        [6].Andco_Values.Pounds_Per_Inch := 65.0, [6].Andco_Values.New_Rate := 4000.0, [6].Andco_Values.Analog := 1, [6].Andco_Values.Min_Position := 625, [6].Andco_Values.Length := 12.0, [6].Andco_Values.InchesOpen := 7.1282053, [6].Andco_Values.AnalogValue := 9660, [6].Clean_Load_Delay_Stop := 36000, [6].Treat_Load_Delay_Stop := 34000, [6].tmrStopDelay.EN := 1, [6].tmrStopDelay.TT := 1, [6].Available_For_Clean_Load := 1, [6].Available_For_Treat_Load := 1, [7].Bin_Description := '10', [7].Bin_Variety.Item_Number := '823001', [7].Bin_Variety.Name := 'ARTDECO CERTIFIED FALL SWH', [7].Bin_Variety.Class := 'Certified', [7].Bin_Variety.Color[0].Color := 1, [7].Rate_Cal_Points[1].Andco_Position := 3007, [7].Rate_Cal_Points[1].Rate := 1000, [7].Rate_Cal_Points[2].Andco_Position := 5443, [7].Rate_Cal_Points[2].Rate := 2000, [7].Rate_Cal_Points[3].Andco_Position := 7342, [7].Rate_Cal_Points[3].Rate := 3000, [7].Rate_Cal_Points[4].Andco_Position := 9304, [7].Rate_Cal_Points[4].Rate := 4000, [7].Clean_Load_Delay_Start := 36500, [7].Treat_Load_Delay_Start := 30000, [7].Andco_Values.Cal_Status := 4, [7].Andco_Values.Raw_Position := 9878, [7].Andco_Values.Max_Position := 10246, [7].Andco_Values.Preact := 20, [7].Andco_Values.Percent_Open := 0.9646484, [7].Andco_Values.New_Pos := 68, [7].Andco_Values.Width := 6.0, [7].Andco_Values.Rate := 4292.5586, [7].Andco_Values.Pounds_Per_Inch := 65.0, [7].Andco_Values.New_Rate := 3700.0, [7].Andco_Values.Analog := 1, [7].Andco_Values.Min_Position := 6, [7].Andco_Values.Length := 12.0, [7].Andco_Values.InchesOpen := 11.575781, [7].Andco_Values.AnalogValue := 9884, [7].Clean_Load_Delay_Stop := 36500, [7].Treat_Load_Delay_Stop := 33000, [7].tmrStopDelay.EN := 1, [7].tmrStopDelay.TT := 1, [7].Available_For_Clean_Load := 1, [7].Available_For_Treat_Load := 1, [8].Bin_Description := '12', [8].Bin_Variety.Name := 'Empty', [8].Bin_Variety.Color[0].Color := 1, [8].Rate_Cal_Points[1].Andco_Position := 3358, [8].Rate_Cal_Points[1].Rate := 1000, [8].Rate_Cal_Points[2].Andco_Position := 5110, [8].Rate_Cal_Points[2].Rate := 2000, [8].Rate_Cal_Points[3].Andco_Position := 6534, [8].Rate_Cal_Points[3].Rate := 3000, [8].Rate_Cal_Points[4].Andco_Position := 8210, [8].Rate_Cal_Points[4].Rate := 4000,
        [8].Clean_Load_Delay_Start := 37000, [8].Treat_Load_Delay_Start := 31000, [8].Andco_Values.Cal_Status := 4, [8].Andco_Values.Raw_Position := 8474, [8].Andco_Values.Max_Position := 15055, [8].Andco_Values.Preact := 20, [8].Andco_Values.Percent_Open := 0.66141117, [8].Andco_Values.New_Pos := 61, [8].Andco_Values.Width := 6.0, [8].Andco_Values.Rate := 4157.518, [8].Andco_Values.Pounds_Per_Inch := 65.0, [8].Andco_Values.New_Rate := 3800.0, [8].Andco_Values.Analog := 1, [8].Andco_Values.Min_Position := 2243, [8].Andco_Values.Length := 12.0, [8].Andco_Values.InchesOpen := 7.936934, [8].Andco_Values.AnalogValue := 10717, [8].Clean_Load_Delay_Stop := 37000, [8].Treat_Load_Delay_Stop := 34000, [8].tmrStopDelay.EN := 1, [8].tmrStopDelay.TT := 1, [8].Available_For_Clean_Load := 1, [8].Available_For_Treat_Load := 1, [9].Bin_Description := '14', [9].Bin_Variety.Item_Number := '873002', [9].Bin_Variety.Name := 'HD-307 CERTIFIED HWW', [9].Bin_Variety.Class := 'Certified', [9].Bin_Variety.Color[0].Color := 1, [9].Rate_Cal_Points[1].Andco_Position := 2158, [9].Rate_Cal_Points[1].Rate := 1000, [9].Rate_Cal_Points[2].Andco_Position := 4887, [9].Rate_Cal_Points[2].Rate := 2000, [9].Rate_Cal_Points[3].Andco_Position := 6612, [9].Rate_Cal_Points[3].Rate := 3000, [9].Rate_Cal_Points[4].Andco_Position := 8287, [9].Rate_Cal_Points[4].Rate := 4000, [9].Clean_Load_Delay_Start := 37500, [9].Treat_Load_Delay_Start := 31000, [9].Andco_Values.Raw_Position := 8668, [9].Andco_Values.Max_Position := 13031, [9].Andco_Values.Preact := 20, [9].Andco_Values.Percent_Open := 0.68679184, [9].Andco_Values.Width := 6.0, [9].Andco_Values.Rate := 4227.463, [9].Andco_Values.Pounds_Per_Inch := 65.0, [9].Andco_Values.Analog := 1, [9].Andco_Values.Min_Position := 410, [9].Andco_Values.Length := 12.0, [9].Andco_Values.InchesOpen := 8.241502, [9].Andco_Values.AnalogValue := 9078, [9].Clean_Load_Delay_Stop := 37500, [9].Treat_Load_Delay_Stop := 34000, [9].tmrStopDelay.EN := 1, [9].tmrStopDelay.TT := 1, [9].Available_For_Clean_Load := 1, [9].Available_For_Treat_Load := 1, [10].Bin_Description := '15', [10].Bin_Variety.Item_Number := '873002', [10].Bin_Variety.Name := 'HD-307 CERTIFIED HWW', [10].Bin_Variety.Class := 'Certified',
        [10].Bin_Variety.Color[0].Color := 1, [10].Rate_Cal_Points[1].Andco_Position := 2321, [10].Rate_Cal_Points[1].Rate := 1000, [10].Rate_Cal_Points[2].Andco_Position := 4523, [10].Rate_Cal_Points[2].Rate := 2000, [10].Rate_Cal_Points[3].Andco_Position := 6483, [10].Rate_Cal_Points[3].Rate := 3000, [10].Rate_Cal_Points[4].Andco_Position := 8309, [10].Rate_Cal_Points[4].Rate := 4000, [10].Clean_Load_Delay_Start := 38000, [10].Treat_Load_Delay_Start := 30000, [10].Andco_Values.Cal_Status := 4, [10].Andco_Values.Raw_Position := 8354, [10].Andco_Values.Max_Position := 12922, [10].Andco_Values.Preact := 20, [10].Andco_Values.Percent_Open := 0.6724082, [10].Andco_Values.Width := 6.0, [10].Andco_Values.Rate := 4024.644, [10].Andco_Values.Pounds_Per_Inch := 65.0, [10].Andco_Values.Analog := 1, [10].Andco_Values.Min_Position := 498, [10].Andco_Values.Length := 12.0, [10].Andco_Values.InchesOpen := 8.068899, [10].Andco_Values.AnalogValue := 8852, [10].Clean_Load_Delay_Stop := 38000, [10].Treat_Load_Delay_Stop := 34000, [10].tmrStartDelay.PRE := 2000, [10].tmrStopDelay.PRE := 2000, [10].tmrStopDelay.EN := 1, [10].tmrStopDelay.TT := 1, [10].StartDelayPre := 2000, [10].StopDelayPre := 2000, [10].Available_For_Clean_Load := 1, [10].Available_For_Treat_Load := 1, [11].Bin_Description := '20', [11].Bin_Variety.Item_Number := '873003', [11].Bin_Variety.Name := 'DAYN CERTIFIED HWW', [11].Bin_Variety.Class := 'Certified', [11].Bin_Variety.Color[0].Color := 1, [11].Rate_Cal_Points[1].Andco_Position := 3830, [11].Rate_Cal_Points[1].Rate := 1000, [11].Rate_Cal_Points[2].Andco_Position := 5231, [11].Rate_Cal_Points[2].Rate := 2000, [11].Rate_Cal_Points[3].Andco_Position := 7521, [11].Rate_Cal_Points[3].Rate := 3000, [11].Rate_Cal_Points[4].Andco_Position := 8755, [11].Rate_Cal_Points[4].Rate := 4000, [11].Clean_Load_Delay_Start := 38000, [11].Treat_Load_Delay_Start := 31000, [11].Andco_Values.Cal_Status := 2, [11].Andco_Values.Raw_Position := 8988, [11].Andco_Values.Max_Position := 12959, [11].Andco_Values.Preact := 32, [11].Andco_Values.Percent_Open := 0.72712564, [11].Andco_Values.New_Pos := 78, [11].Andco_Values.Width := 6.0, [11].Andco_Values.Rate := 4188.817, [11].Andco_Values.Pounds_Per_Inch := 65.0, [11].Andco_Values.New_Rate := 4400.0, [11].Andco_Values.Analog := 1,
        [11].Andco_Values.Min_Position := 598, [11].Andco_Values.Length := 12.0, [11].Andco_Values.InchesOpen := 8.725508, [11].Andco_Values.AnalogValue := 9586, [11].Clean_Load_Delay_Stop := 38000, [11].Treat_Load_Delay_Stop := 35000, [11].tmrStopDelay.EN := 1, [11].tmrStopDelay.TT := 1, [11].Available_For_Clean_Load := 1, [11].Available_For_Treat_Load := 1, [12].Bin_Description := '13', [12].Bin_Variety.Item_Number := '823072', [12].Bin_Variety.Name := 'VOODOO CF CERTIFIED FALL SWH', [12].Bin_Variety.Class := 'Certified', [12].Bin_Variety.Color[0].Color := 1, [12].Rate_Cal_Points[1].Andco_Position := 2243, [12].Rate_Cal_Points[1].Rate := 1000, [12].Rate_Cal_Points[2].Andco_Position := 4281, [12].Rate_Cal_Points[2].Rate := 2000, [12].Rate_Cal_Points[3].Andco_Position := 5779, [12].Rate_Cal_Points[3].Rate := 3000, [12].Rate_Cal_Points[4].Andco_Position := 7567, [12].Rate_Cal_Points[4].Rate := 4000, [12].Clean_Load_Delay_Start := 38500, [12].Treat_Load_Delay_Start := 32000, [12].Andco_Values.Cal_Status := 2, [12].Andco_Values.Raw_Position := 7647, [12].Andco_Values.Max_Position := 12088, [12].Andco_Values.Preact := 20, [12].Andco_Values.Percent_Open := 0.6331346, [12].Andco_Values.New_Pos := 36, [12].Andco_Values.Width := 6.0, [12].Andco_Values.Rate := 4044.7427, [12].Andco_Values.Pounds_Per_Inch := 65.0, [12].Andco_Values.New_Rate := 2500.0, [12].Andco_Values.Analog := 1, [12].Andco_Values.Min_Position := 10, [12].Andco_Values.Length := 12.0, [12].Andco_Values.InchesOpen := 7.5976152, [12].Andco_Values.AnalogValue := 7657, [12].Clean_Load_Delay_Stop := 38500, [12].Treat_Load_Delay_Stop := 36000, [12].tmrStopDelay.EN := 1, [12].tmrStopDelay.TT := 1, [12].Available_For_Clean_Load := 1, [12].Available_For_Treat_Load := 1, [13].Bin_Description := '19', [13].Bin_Variety.Name := 'Empty', [13].Bin_Variety.Color[0].Color := 1, [13].Rate_Cal_Points[1].Andco_Position := 1992, [13].Rate_Cal_Points[1].Rate := 1000, [13].Rate_Cal_Points[2].Andco_Position := 3762, [13].Rate_Cal_Points[2].Rate := 2000, [13].Rate_Cal_Points[3].Andco_Position := 5733, [13].Rate_Cal_Points[3].Rate := 3000, [13].Rate_Cal_Points[4].Andco_Position := 7278, [13].Rate_Cal_Points[4].Rate := 4000, [13].Clean_Load_Delay_Start := 38500, [13].Treat_Load_Delay_Start := 33000, [13].Andco_Values.Cal_Status := 4,
        [13].Andco_Values.Raw_Position := 7215, [13].Andco_Values.Max_Position := 14383, [13].Andco_Values.Preact := 20, [13].Andco_Values.Percent_Open := 0.5766925, [13].Andco_Values.Width := 6.0, [13].Andco_Values.Rate := 3959.2231, [13].Andco_Values.Pounds_Per_Inch := 65.0, [13].Andco_Values.Analog := 1, [13].Andco_Values.Min_Position := 1872, [13].Andco_Values.Length := 12.0, [13].Andco_Values.InchesOpen := 6.92031, [13].Andco_Values.AnalogValue := 9087, [13].Clean_Load_Delay_Stop := 38500, [13].Treat_Load_Delay_Stop := 36000, [13].tmrStopDelay.EN := 1, [13].tmrStopDelay.TT := 1, [13].Available_For_Clean_Load := 1, [13].Available_For_Treat_Load := 1, [14].Bin_Description := '19 SIDE', [14].Bin_Variety.Name := 'Empty', [14].Rate_Cal_Points[1].Andco_Position := 10, [14].Rate_Cal_Points[1].Rate := 1000, [14].Rate_Cal_Points[2].Andco_Position := 20, [14].Rate_Cal_Points[2].Rate := 2000, [14].Rate_Cal_Points[3].Andco_Position := 43, [14].Rate_Cal_Points[3].Rate := 3000, [14].Rate_Cal_Points[4].Andco_Position := 5025, [14].Rate_Cal_Points[4].Rate := 4000, [14].Clean_Load_Delay_Start := 9000, [14].Treat_Load_Delay_Start := 9000, [14].Andco_Values.Raw_Position := 9078, [14].Andco_Values.Max_Position := 120, [14].Andco_Values.Preact := 20, [14].Andco_Values.Percent_Open := 75.65, [14].Andco_Values.Width := 6.0, [14].Andco_Values.Rate := 4813.529, [14].Andco_Values.Pounds_Per_Inch := 65.0, [14].Andco_Values.Analog := 1, [14].Andco_Values.Length := 12.0, [14].Andco_Values.InchesOpen := 907.80005, [14].Andco_Values.AnalogValue := 9078, [14].Clean_Load_Delay_Stop := 9000, [14].Treat_Load_Delay_Stop := 9000, [14].tmrStartDelay.PRE := 4000, [14].tmrStopDelay.PRE := 4000, [14].tmrStopDelay.EN := 1, [14].tmrStopDelay.TT := 1, [14].StartDelayPre := 4000, [14].StopDelayPre := 4000, [14].Available_For_Clean_Load := 1, [14].Available_For_Treat_Load := 1, [15].Bin_Description := '13 SIDE', [15].Bin_Variety.Name := 'Empty', [15].Rate_Cal_Points[1].Andco_Position := 10, [15].Rate_Cal_Points[1].Rate := 1000, [15].Rate_Cal_Points[2].Andco_Position := 20, [15].Rate_Cal_Points[2].Rate := 2000, [15].Rate_Cal_Points[3].Andco_Position := 43, [15].Rate_Cal_Points[3].Rate := 3000, [15].Rate_Cal_Points[4].Andco_Position := 6367,
        [15].Rate_Cal_Points[4].Rate := 4000, [15].Clean_Load_Delay_Start := 9000, [15].Treat_Load_Delay_Start := 9000, [15].Andco_Values.Raw_Position := 8852, [15].Andco_Values.Max_Position := 120, [15].Andco_Values.Preact := 20, [15].Andco_Values.Percent_Open := 73.76667, [15].Andco_Values.Width := 6.0, [15].Andco_Values.Rate := 4392.9473, [15].Andco_Values.Pounds_Per_Inch := 65.0, [15].Andco_Values.Analog := 1, [15].Andco_Values.Length := 12.0, [15].Andco_Values.InchesOpen := 885.2001, [15].Andco_Values.AnalogValue := 8852, [15].Clean_Load_Delay_Stop := 9000, [15].Treat_Load_Delay_Stop := 9000, [15].tmrStopDelay.EN := 1, [15].tmrStopDelay.TT := 1, [15].Available_For_Clean_Load := 1, [15].Available_For_Treat_Load := 1, [16].Bin_Description := '11', [16].Bin_Variety.Item_Number := '823098', [16].Bin_Variety.Name := 'RE-DAG COAXIUM - CERTIFIED', [16].Bin_Variety.Class := 'Certified', [16].Bin_Variety.Color[0].Color := 1, [16].Rate_Cal_Points[1].Andco_Position := 4978, [16].Rate_Cal_Points[1].Rate := 1000, [16].Rate_Cal_Points[2].Andco_Position := 8166, [16].Rate_Cal_Points[2].Rate := 2000, [16].Rate_Cal_Points[3].Andco_Position := 10647, [16].Rate_Cal_Points[3].Rate := 3000, [16].Rate_Cal_Points[4].Andco_Position := 14081, [16].Rate_Cal_Points[4].Rate := 4000, [16].Clean_Load_Delay_Start := 27000, [16].Treat_Load_Delay_Start := 11000, [16].Bindicator_Low := 1, [16].Andco_Values.Cal_Status := 4, [16].Andco_Values.Raw_Position := 13887, [16].Andco_Values.Max_Position := 16180, [16].Andco_Values.Preact := 20, [16].Andco_Values.Percent_Open := 0.9065213, [16].Andco_Values.New_Pos := 101, [16].Andco_Values.Width := 6.0, [16].Andco_Values.Rate := 3943.506, [16].Andco_Values.Pounds_Per_Inch := 65.0, [16].Andco_Values.New_Rate := 4000.0, [16].Andco_Values.Analog := 1, [16].Andco_Values.Min_Position := 861, [16].Andco_Values.Length := 12.0, [16].Andco_Values.InchesOpen := 10.878256, [16].Andco_Values.AnalogValue := 14748, [16].Clean_Load_Delay_Stop := 27000, [16].Treat_Load_Delay_Stop := 12000, [16].tmrStopDelay.EN := 1, [16].tmrStopDelay.TT := 1, [16].Available_For_Clean_Load := 1, [16].Available_For_Treat_Load := 1, [17].Bin_Description := '12', [17].Bin_Variety.Item_Number := '843022', [17].Bin_Variety.Name := 'VENOM CERTIFIED DNS',
        [17].Bin_Variety.Class := 'Certified', [17].Bin_Variety.Color[0].Color := 1, [17].Rate_Cal_Points[1].Andco_Position := 5131, [17].Rate_Cal_Points[1].Rate := 1000, [17].Rate_Cal_Points[2].Andco_Position := 7438, [17].Rate_Cal_Points[2].Rate := 2000, [17].Rate_Cal_Points[3].Andco_Position := 10479, [17].Rate_Cal_Points[3].Rate := 3000, [17].Rate_Cal_Points[4].Andco_Position := 14378, [17].Rate_Cal_Points[4].Rate := 4000, [17].Clean_Load_Delay_Start := 18390, [17].Treat_Load_Delay_Start := 10000, [17].Andco_Values.Fully_Open := 1, [17].Andco_Values.Cal_Status := 4, [17].Andco_Values.Raw_Position := 14945, [17].Andco_Values.Max_Position := 15450, [17].Andco_Values.Preact := 55, [17].Andco_Values.Percent_Open := 0.9995318, [17].Andco_Values.New_Pos := 108, [17].Andco_Values.Width := 6.0, [17].Andco_Values.Rate := 4145.422, [17].Andco_Values.Pounds_Per_Inch := 65.0, [17].Andco_Values.New_Rate := 4000.0, [17].Andco_Values.Analog := 1, [17].Andco_Values.Min_Position := 498, [17].Andco_Values.Length := 12.0, [17].Andco_Values.InchesOpen := 11.994382, [17].Andco_Values.AnalogValue := 15443, [17].Clean_Load_Delay_Stop := 18390, [17].Treat_Load_Delay_Stop := 11000, [17].tmrStopDelay.EN := 1, [17].tmrStopDelay.TT := 1, [17].Available_For_Clean_Load := 1, [17].Available_For_Treat_Load := 1, [18].Bin_Description := '13', [18].Bin_Variety.Name := 'Empty', [18].Bin_Variety.Color[0].Color := 1, [18].Rate_Cal_Points[1].Andco_Position := 4915, [18].Rate_Cal_Points[1].Rate := 1000, [18].Rate_Cal_Points[2].Andco_Position := 7628, [18].Rate_Cal_Points[2].Rate := 2000, [18].Rate_Cal_Points[3].Andco_Position := 12268, [18].Rate_Cal_Points[3].Rate := 3000, [18].Rate_Cal_Points[4].Andco_Position := 13372, [18].Rate_Cal_Points[4].Rate := 4000, [18].Clean_Load_Delay_Start := 17440, [18].Treat_Load_Delay_Start := 10000, [18].Andco_Values.Cal_Status := 2, [18].Andco_Values.Raw_Position := 13995, [18].Andco_Values.Max_Position := 16053, [18].Andco_Values.Preact := 20, [18].Andco_Values.Percent_Open := 0.8855353, [18].Andco_Values.Width := 6.0, [18].Andco_Values.Rate := 4564.3115, [18].Andco_Values.Pounds_Per_Inch := 65.0, [18].Andco_Values.Analog := 1, [18].Andco_Values.Min_Position := 249, [18].Andco_Values.Length := 12.0, [18].Andco_Values.InchesOpen := 10.626424, [18].Andco_Values.AnalogValue := 14244,
        [18].Treat_Load_Delay_Stop := 11000, [18].tmrStopDelay.EN := 1, [18].tmrStopDelay.TT := 1, [18].Available_For_Clean_Load := 1, [18].Available_For_Treat_Load := 1, [19].Bin_Description := '14', [19].Bin_Variety.Item_Number := '822087', [19].Bin_Variety.Name := 'LCS ECLIPSE AX - 0225 COAXIUM REGISTERED HRW', [19].Bin_Variety.Class := 'Registered', [19].Bin_Variety.Color[0].Color := 1, [19].Rate_Cal_Points[1].Andco_Position := 3696, [19].Rate_Cal_Points[1].Rate := 1000, [19].Rate_Cal_Points[2].Andco_Position := 6573, [19].Rate_Cal_Points[2].Rate := 2000, [19].Rate_Cal_Points[3].Andco_Position := 9630, [19].Rate_Cal_Points[3].Rate := 3000, [19].Rate_Cal_Points[4].Andco_Position := 12560, [19].Rate_Cal_Points[4].Rate := 4000, [19].Clean_Load_Delay_Start := 16610, [19].Treat_Load_Delay_Start := 10000, [19].Andco_Values.Cal_Status := 4, [19].Andco_Values.Raw_Position := 12753, [19].Andco_Values.Max_Position := 16151, [19].Andco_Values.Preact := 20, [19].Andco_Values.Percent_Open := 0.8254369, [19].Andco_Values.Width := 6.0, [19].Andco_Values.Rate := 4065.8704, [19].Andco_Values.Pounds_Per_Inch := 65.0, [19].Andco_Values.Analog := 1, [19].Andco_Values.Min_Position := 701, [19].Andco_Values.Length := 12.0, [19].Andco_Values.InchesOpen := 9.905243, [19].Andco_Values.AnalogValue := 13454, [19].Clean_Load_Delay_Stop := 16610, [19].Treat_Load_Delay_Stop := 9000, [19].tmrStopDelay.EN := 1, [19].tmrStopDelay.TT := 1, [19].Available_For_Clean_Load := 1, [19].Available_For_Treat_Load := 1, [20].Bin_Description := '15', [20].Bin_Variety.Item_Number := '803003', [20].Bin_Variety.Name := 'JET CERTIFIED HRW', [20].Bin_Variety.Class := 'Certified', [20].Bin_Variety.Color[0].Color := 1, [20].Rate_Cal_Points[1].Andco_Position := 4509, [20].Rate_Cal_Points[1].Rate := 1000, [20].Rate_Cal_Points[2].Andco_Position := 7812, [20].Rate_Cal_Points[2].Rate := 2000, [20].Rate_Cal_Points[3].Andco_Position := 10414, [20].Rate_Cal_Points[3].Rate := 3000, [20].Rate_Cal_Points[4].Andco_Position := 13301, [20].Rate_Cal_Points[4].Rate := 4000, [20].Clean_Load_Delay_Start := 15870, [20].Treat_Load_Delay_Start := 9000, [20].Andco_Values.Cal_Status := 4, [20].Andco_Values.Raw_Position := 14405, [20].Andco_Values.Max_Position := 15728, [20].Andco_Values.Preact := 20, [20].Andco_Values.Percent_Open := 0.9190965, [20].Andco_Values.New_Pos := 7461,
        [20].Andco_Values.Width := 6.0, [20].Andco_Values.Rate := 4382.404, [20].Andco_Values.Pounds_Per_Inch := 65.0, [20].Andco_Values.New_Rate := 3800.0, [20].Andco_Values.Analog := 1, [20].Andco_Values.Min_Position := 55, [20].Andco_Values.Length := 12.0, [20].Andco_Values.InchesOpen := 11.029159, [20].Andco_Values.AnalogValue := 14460, [20].Treat_Load_Delay_Stop := 9000, [20].tmrStopDelay.EN := 1, [20].tmrStopDelay.TT := 1, [20].Available_For_Clean_Load := 1, [20].Available_For_Treat_Load := 1, [21].Bin_Description := '16', [21].Bin_Variety.Item_Number := '823093', [21].Bin_Variety.Name := 'SCORPION COAX-0291 CERTIFIED SWH', [21].Bin_Variety.Class := 'Certified', [21].Bin_Variety.Color[0].Color := 1, [21].Rate_Cal_Points[1].Andco_Position := 5171, [21].Rate_Cal_Points[1].Rate := 1000, [21].Rate_Cal_Points[2].Andco_Position := 8208, [21].Rate_Cal_Points[2].Rate := 2000, [21].Rate_Cal_Points[3].Andco_Position := 11698, [21].Rate_Cal_Points[3].Rate := 3000, [21].Rate_Cal_Points[4].Andco_Position := 14346, [21].Rate_Cal_Points[4].Rate := 4000, [21].Clean_Load_Delay_Start := 19000, [21].Treat_Load_Delay_Start := 8000, [21].Bindicator_Low := 1, [21].Andco_Values.Cal_Status := 4, [21].Andco_Values.Raw_Position := 5924, [21].Andco_Values.Max_Position := 16315, [21].Andco_Values.Preact := 20, [21].Andco_Values.Percent_Open := 0.37267238, [21].Andco_Values.New_Pos := 133, [21].Andco_Values.Width := 6.0, [21].Andco_Values.Rate := 1247.942, [21].Andco_Values.Pounds_Per_Inch := 65.0, [21].Andco_Values.New_Rate := 5000.0, [21].Andco_Values.Analog := 1, [21].Andco_Values.Min_Position := 419, [21].Andco_Values.Length := 12.0, [21].Andco_Values.InchesOpen := 4.472069, [21].Andco_Values.AnalogValue := 6343, [21].Clean_Load_Delay_Stop := 19000, [21].Treat_Load_Delay_Stop := 9000, [21].tmrStartDelay.PRE := 21000, [21].tmrStopDelay.PRE := 23000, [21].tmrStopDelay.EN := 1, [21].tmrStopDelay.TT := 1, [21].StartDelayPre := 21000, [21].StopDelayPre := 23000, [21].Available_For_Clean_Load := 1, [21].Available_For_Treat_Load := 1, [22].Bin_Description := '17', [22].Bin_Variety.Item_Number := '843036', [22].Bin_Variety.Name := 'HALE CERTIFIED DNS', [22].Bin_Variety.Class := 'Certified', [22].Bin_Variety.Color[0].Color := 1,
        [22].Rate_Cal_Points[1].Andco_Position := 1803, [22].Rate_Cal_Points[1].Rate := 1000, [22].Rate_Cal_Points[2].Andco_Position := 3716, [22].Rate_Cal_Points[2].Rate := 2000, [22].Rate_Cal_Points[3].Andco_Position := 5315, [22].Rate_Cal_Points[3].Rate := 3000, [22].Rate_Cal_Points[4].Andco_Position := 7606, [22].Rate_Cal_Points[4].Rate := 4000, [22].Clean_Load_Delay_Start := 19000, [22].Treat_Load_Delay_Start := 7000, [22].Bindicator_Low := 1, [22].Andco_Values.Cal_Status := 4, [22].Andco_Values.Raw_Position := 7779, [22].Andco_Values.Max_Position := 15450, [22].Andco_Values.Preact := 20, [22].Andco_Values.Percent_Open := 0.5375579, [22].Andco_Values.New_Pos := 47, [22].Andco_Values.Width := 6.0, [22].Andco_Values.Rate := 4075.513, [22].Andco_Values.Pounds_Per_Inch := 65.0, [22].Andco_Values.New_Rate := 4000.0, [22].Andco_Values.Analog := 1, [22].Andco_Values.Min_Position := 979, [22].Andco_Values.Length := 12.0, [22].Andco_Values.InchesOpen := 6.450695, [22].Andco_Values.AnalogValue := 8758, [22].Clean_Load_Delay_Stop := 19000, [22].Treat_Load_Delay_Stop := 10000, [22].tmrStartDelay.PRE := 23000, [22].tmrStopDelay.PRE := 23000, [22].tmrStopDelay.EN := 1, [22].tmrStopDelay.TT := 1, [22].StartDelayPre := 23000, [22].StopDelayPre := 23000, [22].Available_For_Clean_Load := 1, [22].Available_For_Treat_Load := 1, [23].Bin_Description := '21', [23].Bin_Variety.Item_Number := '843001', [23].Bin_Variety.Name := 'BUCK PRONTO CERTIFIED DNS', [23].Bin_Variety.Class := 'Certified', [23].Bin_Variety.Color[0].Color := 1, [23].Rate_Cal_Points[1].Andco_Position := 5036, [23].Rate_Cal_Points[1].Rate := 1000, [23].Rate_Cal_Points[2].Andco_Position := 8241, [23].Rate_Cal_Points[2].Rate := 2000, [23].Rate_Cal_Points[3].Andco_Position := 12245, [23].Rate_Cal_Points[3].Rate := 3000, [23].Rate_Cal_Points[4].Andco_Position := 14788, [23].Rate_Cal_Points[4].Rate := 4000, [23].Clean_Load_Delay_Start := 19000, [23].Treat_Load_Delay_Start := 11000, [23].Bindicator_Low := 1, [23].Andco_Values.Cal_Status := 4, [23].Andco_Values.Raw_Position := 15207, [23].Andco_Values.Max_Position := 16384, [23].Andco_Values.Preact := 20, [23].Andco_Values.Percent_Open := 0.9718796, [23].Andco_Values.New_Pos := 86, [23].Andco_Values.Width := 6.0, [23].Andco_Values.Rate := 4164.766,
        [23].Andco_Values.Pounds_Per_Inch := 65.0, [23].Andco_Values.New_Rate := 4000.0, [23].Andco_Values.Analog := 1, [23].Andco_Values.Min_Position := 737, [23].Andco_Values.Length := 12.0, [23].Andco_Values.InchesOpen := 11.662556, [23].Andco_Values.AnalogValue := 15944, [23].Clean_Load_Delay_Stop := 19000, [23].Treat_Load_Delay_Stop := 14000, [23].tmrStopDelay.EN := 1, [23].tmrStopDelay.TT := 1, [23].Available_For_Clean_Load := 1, [23].Available_For_Treat_Load := 1, [24].Bin_Description := '22', [24].Bin_Variety.Item_Number := '843002', [24].Bin_Variety.Name := 'EXPRESSO CERTIFIED DNS', [24].Bin_Variety.Class := 'Certified', [24].Bin_Variety.Color[0].Color := 1, [24].Rate_Cal_Points[1].Andco_Position := 5147, [24].Rate_Cal_Points[1].Rate := 1000, [24].Rate_Cal_Points[2].Andco_Position := 8427, [24].Rate_Cal_Points[2].Rate := 2000, [24].Rate_Cal_Points[3].Andco_Position := 12356, [24].Rate_Cal_Points[3].Rate := 3000, [24].Rate_Cal_Points[4].Andco_Position := 14863, [24].Rate_Cal_Points[4].Rate := 4000, [24].Clean_Load_Delay_Start := 23500, [24].Treat_Load_Delay_Start := 14000, [24].Bindicator_Low := 1, [24].Andco_Values.Cal_Status := 4, [24].Andco_Values.Raw_Position := 14817, [24].Andco_Values.Max_Position := 16384, [24].Andco_Values.Preact := 20, [24].Andco_Values.Percent_Open := 0.9250796, [24].Andco_Values.New_Pos := 57, [24].Andco_Values.Width := 6.0, [24].Andco_Values.Rate := 3981.6514, [24].Andco_Values.Pounds_Per_Inch := 65.0, [24].Andco_Values.New_Rate := 2000.0, [24].Andco_Values.Analog := 1, [24].Andco_Values.Min_Position := 367, [24].Andco_Values.Length := 12.0, [24].Andco_Values.InchesOpen := 11.100955, [24].Andco_Values.AnalogValue := 15184, [24].Clean_Load_Delay_Stop := 23500, [24].Treat_Load_Delay_Stop := 15000, [24].tmrStartDelay.PRE := 15000, [24].tmrStopDelay.PRE := 17000, [24].tmrStopDelay.EN := 1, [24].tmrStopDelay.TT := 1, [24].StartDelayPre := 15000, [24].StopDelayPre := 17000, [24].Available_For_Clean_Load := 1, [24].Available_For_Treat_Load := 1, [25].Bin_Description := '23', [25].Bin_Variety.Item_Number := '843022', [25].Bin_Variety.Name := 'VENOM CERTIFIED DNS', [25].Bin_Variety.Class := 'Certified', [25].Rate_Cal_Points[1].Andco_Position := 4846, [25].Rate_Cal_Points[1].Rate := 1000,
        [25].Rate_Cal_Points[2].Andco_Position := 8120, [25].Rate_Cal_Points[2].Rate := 2000, [25].Rate_Cal_Points[3].Andco_Position := 11636, [25].Rate_Cal_Points[3].Rate := 3000, [25].Rate_Cal_Points[4].Andco_Position := 13864, [25].Rate_Cal_Points[4].Rate := 4000, [25].Clean_Load_Delay_Start := 28000, [25].Treat_Load_Delay_Start := 18000, [25].Bindicator_Low := 1, [25].Andco_Values.Cal_Status := 4, [25].Andco_Values.Raw_Position := 14906, [25].Andco_Values.Max_Position := 16033, [25].Andco_Values.Preact := 20, [25].Andco_Values.Percent_Open := 0.9807869, [25].Andco_Values.New_Pos := 8762, [25].Andco_Values.Width := 6.0, [25].Andco_Values.Rate := 4467.684, [25].Andco_Values.Pounds_Per_Inch := 65.0, [25].Andco_Values.New_Rate := 3800.0, [25].Andco_Values.Analog := 1, [25].Andco_Values.Min_Position := 835, [25].Andco_Values.Length := 12.0, [25].Andco_Values.InchesOpen := 11.7694435, [25].Andco_Values.AnalogValue := 15741, [25].Clean_Load_Delay_Stop := 28000, [25].Treat_Load_Delay_Stop := 20000, [25].tmrStopDelay.EN := 1, [25].tmrStopDelay.TT := 1, [25].Available_For_Clean_Load := 1, [25].Available_For_Treat_Load := 1, [26].Bin_Description := '24', [26].Bin_Variety.Item_Number := '803003', [26].Bin_Variety.Name := 'JET CERTIFIED HRW', [26].Bin_Variety.Class := 'Certified', [26].Bin_Variety.Color[0].Color := 1, [26].Rate_Cal_Points[1].Andco_Position := 5096, [26].Rate_Cal_Points[1].Rate := 1000, [26].Rate_Cal_Points[2].Andco_Position := 8425, [26].Rate_Cal_Points[2].Rate := 2000, [26].Rate_Cal_Points[3].Andco_Position := 12377, [26].Rate_Cal_Points[3].Rate := 3000, [26].Rate_Cal_Points[4].Andco_Position := 14785, [26].Rate_Cal_Points[4].Rate := 4000, [26].Clean_Load_Delay_Start := 23000, [26].Treat_Load_Delay_Start := 16000, [26].Andco_Values.Cal_Status := 4, [26].Andco_Values.Raw_Position := 14844, [26].Andco_Values.Max_Position := 16384, [26].Andco_Values.Preact := 20, [26].Andco_Values.Percent_Open := 0.93071663, [26].Andco_Values.New_Pos := 76, [26].Andco_Values.Width := 6.0, [26].Andco_Values.Rate := 4024.5017, [26].Andco_Values.Pounds_Per_Inch := 65.0, [26].Andco_Values.New_Rate := 3800.0, [26].Andco_Values.Analog := 1, [26].Andco_Values.Min_Position := 435, [26].Andco_Values.Length := 12.0, [26].Andco_Values.InchesOpen := 11.1686, [26].Andco_Values.AnalogValue := 15279,
        [26].Clean_Load_Delay_Stop := 23000, [26].Treat_Load_Delay_Stop := 16000, [26].tmrStartDelay.PRE := 5000, [26].tmrStopDelay.PRE := 8000, [26].tmrStopDelay.EN := 1, [26].tmrStopDelay.TT := 1, [26].StartDelayPre := 5000, [26].StopDelayPre := 8000, [26].Available_For_Clean_Load := 1, [26].Available_For_Treat_Load := 1, [27].Bin_Description := '25', [27].Bin_Variety.Item_Number := '823087', [27].Bin_Variety.Name := 'LCS ECLIPSE AX - 0225 COAXIUM CERTIFIED HRW', [27].Bin_Variety.Class := 'Certified', [27].Bin_Variety.Color[0].Color := 1, [27].Rate_Cal_Points[1].Andco_Position := 5099, [27].Rate_Cal_Points[1].Rate := 1000, [27].Rate_Cal_Points[2].Andco_Position := 8615, [27].Rate_Cal_Points[2].Rate := 2000, [27].Rate_Cal_Points[3].Andco_Position := 12478, [27].Rate_Cal_Points[3].Rate := 3000, [27].Rate_Cal_Points[4].Andco_Position := 14424, [27].Rate_Cal_Points[4].Rate := 4000, [27].Clean_Load_Delay_Start := 27000, [27].Treat_Load_Delay_Start := 17000, [27].Bindicator_Low := 1, [27].Andco_Values.Cal_Status := 4, [27].Andco_Values.Raw_Position := 14595, [27].Andco_Values.Max_Position := 16121, [27].Andco_Values.Preact := 20, [27].Andco_Values.Percent_Open := 0.9062403, [27].Andco_Values.Width := 6.0, [27].Andco_Values.Rate := 4087.8726, [27].Andco_Values.Pounds_Per_Inch := 65.0, [27].Andco_Values.Analog := 1, [27].Andco_Values.Min_Position := 16, [27].Andco_Values.Length := 12.0, [27].Andco_Values.InchesOpen := 10.874884, [27].Andco_Values.AnalogValue := 14611, [27].Clean_Load_Delay_Stop := 27000, [27].Treat_Load_Delay_Stop := 21000, [27].tmrStopDelay.EN := 1, [27].tmrStopDelay.TT := 1, [27].Available_For_Clean_Load := 1, [27].Available_For_Treat_Load := 1, [28].Bin_Description := '26', [28].Bin_Variety.Item_Number := '803021', [28].Bin_Variety.Name := 'LCS BLACKBIRD CERTIFIED HRW', [28].Bin_Variety.Class := 'Certified', [28].Bin_Variety.Color[0].Color := 1, [28].Rate_Cal_Points[1].Andco_Position := 3558, [28].Rate_Cal_Points[1].Rate := 1000, [28].Rate_Cal_Points[2].Andco_Position := 7029, [28].Rate_Cal_Points[2].Rate := 2000, [28].Rate_Cal_Points[3].Andco_Position := 10092, [28].Rate_Cal_Points[3].Rate := 3000, [28].Rate_Cal_Points[4].Andco_Position := 13120, [28].Rate_Cal_Points[4].Rate := 4000, [28].Clean_Load_Delay_Start := 31000, [28].Treat_Load_Delay_Start := 21000,
        [28].Bindicator_Low := 1, [28].Andco_Values.Cal_Status := 4, [28].Andco_Values.Raw_Position := 15129, [28].Andco_Values.Max_Position := 15233, [28].Andco_Values.Preact := 20, [28].Andco_Values.Percent_Open := 0.994217, [28].Andco_Values.New_Pos := 95, [28].Andco_Values.Width := 6.0, [28].Andco_Values.Rate := 4663.474, [28].Andco_Values.Pounds_Per_Inch := 65.0, [28].Andco_Values.New_Rate := 3800.0, [28].Andco_Values.Analog := 1, [28].Andco_Values.Min_Position := 16, [28].Andco_Values.Length := 12.0, [28].Andco_Values.InchesOpen := 11.930604, [28].Andco_Values.AnalogValue := 15145, [28].Clean_Load_Delay_Stop := 31000, [28].Treat_Load_Delay_Stop := 24000, [28].tmrStopDelay.EN := 1, [28].tmrStopDelay.TT := 1, [28].Available_For_Clean_Load := 1, [28].Available_For_Treat_Load := 1);
   Loadout_K_Valve : udt_Loadout_K_Valve[2] := ([0].Clean_Gate_Opened := 1, [1].Clean_Gate_Opened := 1);
   Loadout_K_Valve_Control : Loadout_K_Valve_Control[2];
   Loadout_KValve_Not_Used : BOOL;
   Longest_Clean_IDX : DINT := 21;
   Longest_Clean_Start_IDX : DINT;
   Longest_Clean_Start_Time : DINT;
   Longest_Clean_Stop_IDX : DINT;
   Longest_Clean_Stop_Time : DINT;
   Longest_Clean_Time : DINT;
   Longest_IDX : DINT := 5;
   Longest_Time : DINT := 60000;
   Longest_Time_IDX : DINT;
   Longest_Treat_IDX : DINT;
   Longest_Treat_Start_IDX : DINT;
   Longest_Treat_Start_Time : DINT;
   Longest_Treat_Stop_IDX : DINT;
   Longest_Treat_Stop_Time : DINT;
   Longest_Treat_Time : DINT;
   Loop_Idx : DINT := 14;
   Man_Start_Stop_Allowed : BOOL := 1;
   Manual_Blow_Out : BOOL;
   Manual_Mode : BOOL;
   Manual_Open_Calibration_Valves : BOOL;
   Manually_Start_Treater : BOOL;
   Move_Bin_Config : BOOL;
   NA : BOOL;
   New_DeltaX : REAL := -23.0;
   New_DeltaY : REAL := -1000.0;
   Ok_Stop_Belt : BOOL;
   Open_Clean_Bins : BOOL;
   Open_Transfer_Bins : BOOL;
   Open_Treat_Bins : BOOL;
   Pause_Load : BOOL;
   Pause_Load_By_Time : BOOL[32];
   Pause_Load_By_Weight : BOOL[32];
   Pause_Load_Expired : DINT[2];
   Pause_Load_Pre : DINT[2] := ([0] := 29000, [1] := 32000);
   Pause_Transfer_By_Time : BOOL;
   Pause_Transfer_Load_Expired : DINT;
   Pause_Transfer_Msc : DINT := 1800000;
   Pause_Transfer_Pre : DINT := 30;
   Pause_Treat_By_Time : BOOL;
   Pause_Treat_Pre : DINT;
   Pause_Treatment : BOOL;
   Point1 : DINT := 3;
   Point2 : DINT := 4;
   Probe_Above_K_Valve : BOOL;
   Produced_Motor_Values : DINT;
   Rate_Mult : REAL := 0.33025098;
   Remote_Pause_Treat : BOOL;
   Request_Variety : udt_Requested_Variety := (Item_Number := '123', Percentage := 1.0, Bin_Available := 1);
   Requested_Varieties : udt_Requested_Variety[10] := ([0].Item_Number := '123456', [0].Percentage := 0.5, [0].Bin_Available := 1);
   Reset_Bin_Cal : BOOL := 1;
   Reset_Remote_Pause : BOOL;
   Reset_Treat_Chemicals : BOOL;
   ResetSelectedBins : BOOL := 1;
   Rev_Delay_Latch_FWD : BOOL;
   Rev_Delay_Latch_REV : BOOL;
   Reverse_Belt_Forward_Interlock : BOOL := 1;
   Reverse_Belt_Stopping : BOOL;
   Reversing_Belt_Bypass_Valve : BOOL := 1;
   Reversing_Belt_Fans : udt_Cyclone;
   Reversing_Belt_Name : STRING; {constant}
   Reversing_Belt_Reversed : BOOL;
   Scale : SCALE;
   Scale_Target : DINT;
   SCL_01 : SCALE;
   SCL_02 : SCALE;
   SCL_03 : SCALE;
   SCL_04 : SCALE;
   SCL_05 : SCALE;
   SCL_06 : SCALE;
   SCL_07 : SCALE;
   SCL_08 : SCALE := (InRawMax := 30000.0, InEUMax := 50.0);
   SCL_16 : SCALE := (In := 3976.0, InRawMax := 20000.0, InRawMin := 4000.0, InEUMax := 200.0, Out := -0.3, MinAlarm := 1);
   SCL_AMP_Belt10 : SCALE := (In := 10.0, InRawMax := 30151.0, InEUMax := 50.0, Out := 0.016583197);
   SCL_AMP_Belt11 : SCALE := (In := -1.0, InRawMax := 30154.0, InEUMax := 50.0, Out := -0.0016581548, MinAlarm := 1);
   SCL_AMP_Belt11_01 : SCALE;
   SCL_AMP_Belt7 : SCALE := (In := -53.0, InRawMax := 41874.0, InEUMax := 200.0, Out := -0.2531404, MinAlarm := 1);
   SCL_AMP_Belt7_01 : SCALE;
   SCL_AMP_Belt8 : SCALE := (In := 1.0, InRawMax := 29984.0, InEUMax := 50.0, Out := 0.001667556);
   SCL_AMP_Belt8_01 : SCALE;
   SCL_AMP_Belt9 : SCALE := (In := 18.0, InRawMax := 30000.0, InEUMax := 50.0, Out := 0.030000001);
   SCL_AMP_BIN16_AUG : SCALE := (InRawMax := 30000.0, InEUMax := 50.0);
   SCL_AMP_Bin17_AUG : SCALE;
   SCL_AMPS_Belt4 : SCALE := (In := -11.0, InRawMax := 41623.0, InEUMax := 200.0, Out := -0.05285539, MinAlarm := 1);
   SCL_AMPS_Belt5 : SCALE := (In := 11.0, InRawMax := 30168.0, InEUMax := 50.0, Out := 0.018231237);
   SCL_AMPS_Belt6 : SCALE := (In := 8.0, InRawMax := 30203.0, InEUMax := 50.0, Out := 0.013243717);
   Select_Bin_Load_Type : DINT;
   Select_Bin_To_Cal : BOOL;
   Slope : REAL := 1.992;
   Sort_Time_Idx : DINT;
   Sorted_Times : DINT[29,2];
   Start_Bin_Cal : BOOL;
   Start_Blower_707 : BOOL;
   Start_Clean_Belts_Enabled : BOOL;
   Start_Rev_Mtr : udt_Motor_Start;
   Start_Treat_Belts_Enabled : BOOL;
   Steel_Bin_Timing_Offset : DINT := -5;
   Steel_Rqd_Belts_Running : BOOL;
   Stop_Treater : BOOL;
   SUBTest1 : DINT;
   SubTest2 : DINT;
   System_In_Use : BOOL;
   System_Status_Msg : STRING := 'System$0D$0AIdle';
   System_Status_Msgs : STRING[20] := ([0] := 'System$0D$0AIdle', [1] := 'Manual Mode$0D$0A NO INTERLOCKS ! $0D$0A (Be Careful)');
   Target_Weight : DINT[2] := ([0] := 18800, [1] := 78000);
   Test1 : BOOL;
   Test_10Slp : BOOL;
   Test_20Slp : BOOL := 1;
   Test_Air_Gate : BOOL;
   Test_Air_Gate25 : BOOL;
   Test_Air_Open_Input : BOOL;
   Test_In : BOOL;
   Test_Int : DINT;
   Test_Plug : BOOL;
   TestAmps : DINT;
   TestReal : REAL := 1.235;
   Time_Sorter : CONTROL := (LEN := 29);
   Timed_Gate_Met : DINT;
   Timer_Target : REAL;
   tmr_Auto_Start : TIMER := (PRE := 1000, ACC := 1005);
   tmr_Blow_Out : TIMER := (ACC := 16, EN := 1, DN := 1);
   TMR_Concrete_Fan : TIMER := (PRE := 180000, ACC := 180014);
   TMR_Max_Clean_Delay : TIMER;
   TMR_Max_Treat_Delay : TIMER;
   tmr_Pause_Load_Timer : TIMER[2] := ([0].PRE := 29000, [1].PRE := 32000);
   tmr_Pause_Transfer_Timer : TIMER := (PRE := 1800000);
   tmr_Pause_Treat_Timer : TIMER;
   TMR_Reverse_Delay : TIMER := (PRE := 4000, ACC := 4001);
   tmr_Setpoint : TIMER;
   tmrBin_Delay_Start : TIMER[30] := ([0].PRE := 10000, [0].ACC := 10008, [0].EN := 1, [0].DN := 1, [1].PRE := 5000);
   tmrCleanSetpoint : TIMER;
   tmrCleanTime : TIMER := (PRE := 1000);
   tmrDelayTreatStart : TIMER := (PRE := 30000);
   tmrDelayTreatStop : TIMER := (PRE := 33000);
   tmrResetChemicals : TIMER := (PRE := 1000);
   tmrTransferTime : TIMER := (PRE := 1000);
   tmrTreatSetpoint : TIMER;
   tmrTreatTime : TIMER := (PRE := 1000);
   Transfer_Batch_Status : DINT;
   Transfer_Belts_Starting : BOOL;
   Transfer_From_IDX : DINT := -1;
   Transfer_Interlock : BOOL;
   Transfer_To_IDX : DINT := -1;
   TransferHours : DINT;
   TransferMinuets : DINT;
   TransferSeconds : DINT;
   Treat_Batch_Status : DINT;
   Treat_Bin_Gates_Opened : BOOL := 1;
   Treat_Bins_Open : BOOL;
   Treat_Bins_Ready : BOOL := 1;
   Treat_Interlock : BOOL;
   Treat_Jump_Interlock : BOOL;
   Treat_Load : BOOL;
   Treat_Scale_Target : DINT;
   Treat_Scale_Unavailable : BOOL;
   Treater_Calibration : BOOL;
   Treater_Loadout : udt_Treater_Loadout := (Use_A_Treater := 1, Use_B_Treater := 1, Drip_Gate_Closed := 1);
   Treater_Loadout_Open_Bins : BOOL;
   TreatHours : DINT;
   Treatment_Running : BOOL;
   Treatment_Started : BOOL;
   TreatMinuets : DINT;
   TreatSeconds : DINT;
   Truck_Scale_Control : Truck_Scale_Control[3];
   Use_Concrete_Side_Clean : BOOL;
   Use_Concrete_Side_Treat : BOOL;
   Use_Steel_Side_Clean : BOOL;
   Use_Steel_Side_Treat : BOOL;
   Use_Steel_Transfer_Bins : BOOL;
   X1 : REAL;
   X2 : REAL := 1000.0;
   Y1 : REAL;
   Y2 : REAL := 1992.0;
   ZZTEST : udt_Motor_Start;
END_VAR
